// TIA Portal project "OpenLibraryExample" (V13) (continued)
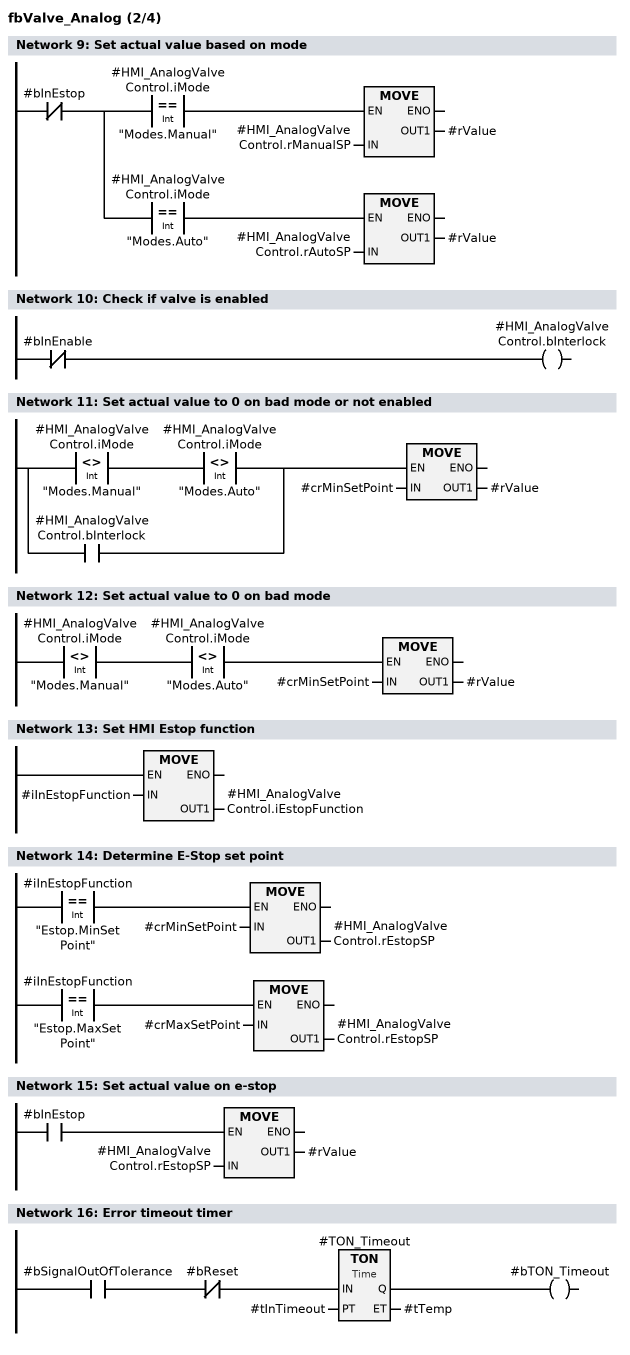
   RUNG wire#powerrail
      I_Contact( #bInEstop )
      wire#w1
      { S7_Templates := "SrcType := Int" } EQ_Contact(in1 := #HMI_AnalogValveControl.iMode, in2 := "Modes.Manual")
      { S7_GenerateENO := "TRUE" } Move(in := #HMI_AnalogValveControl.rManualSP, out1 => #rValue)
   END_RUNG
   RUNG wire#w1
      { S7_Templates := "SrcType := Int" } EQ_Contact(in1 := #HMI_AnalogValveControl.iMode, in2 := "Modes.Auto")
      { S7_GenerateENO := "TRUE" } Move(in := #HMI_AnalogValveControl.rAutoSP, out1 => #rValue)
   END_RUNG
   // the same network as SCL:
   IF NOT #bInEstop AND (#HMI_AnalogValveControl.iMode = "Modes.Manual") THEN
       #rValue := #HMI_AnalogValveControl.rManualSP;
   END_IF;
   IF NOT #bInEstop AND (#HMI_AnalogValveControl.iMode = "Modes.Auto") THEN
       #rValue := #HMI_AnalogValveControl.rAutoSP;
   END_IF;
END_REGION

REGION Network 10: Check if valve is enabled
   RUNG wire#powerrail
      I_Contact( #bInEnable )
      Coil( #HMI_AnalogValveControl.bInterlock )
   END_RUNG
   // the same network as SCL:
   #HMI_AnalogValveControl.bInterlock := NOT #bInEnable;
END_REGION

REGION Network 11: Set actual value to 0 on bad mode or not enabled
   RUNG wire#powerrail
      { S7_Templates := "SrcType := Int" } NE_Contact(in1 := #HMI_AnalogValveControl.iMode, in2 := "Modes.Manual")
      { S7_Templates := "SrcType := Int" } NE_Contact(in1 := #HMI_AnalogValveControl.iMode, in2 := "Modes.Auto")
      wire#w1
      { S7_GenerateENO := "TRUE" } Move(in := #crMinSetPoint, out1 => #rValue)
   END_RUNG
   RUNG wire#powerrail
      Contact( #HMI_AnalogValveControl.bInterlock )
   END_RUNG wire#w1
   // the same network as SCL:
   IF ((#HMI_AnalogValveControl.iMode <> "Modes.Manual") AND (#HMI_AnalogValveControl.iMode <> "Modes.Auto")) OR #HMI_AnalogValveControl.bInterlock THEN
       #rValue := #crMinSetPoint;
   END_IF;
END_REGION

REGION Network 12: Set actual value to 0 on bad mode
   RUNG wire#powerrail
      { S7_Templates := "SrcType := Int" } NE_Contact(in1 := #HMI_AnalogValveControl.iMode, in2 := "Modes.Manual")
      { S7_Templates := "SrcType := Int" } NE_Contact(in1 := #HMI_AnalogValveControl.iMode, in2 := "Modes.Auto")
      { S7_GenerateENO := "TRUE" } Move(in := #crMinSetPoint, out1 => #rValue)
   END_RUNG
   // the same network as SCL:
   IF (#HMI_AnalogValveControl.iMode <> "Modes.Manual") AND (#HMI_AnalogValveControl.iMode <> "Modes.Auto") THEN
       #rValue := #crMinSetPoint;
   END_IF;
END_REGION

REGION Network 13: Set HMI Estop function
   RUNG wire#powerrail
      Move(in := #iInEstopFunction, out1 => #HMI_AnalogValveControl.iEstopFunction)
   END_RUNG
   // the same network as SCL:
   #HMI_AnalogValveControl.iEstopFunction := #iInEstopFunction;
END_REGION

REGION Network 14: Determine E-Stop set point
   RUNG wire#powerrail
      { S7_Templates := "SrcType := Int" } EQ_Contact(in1 := #iInEstopFunction, in2 := "Estop.MinSetPoint")
      { S7_GenerateENO := "TRUE" } Move(in := #crMinSetPoint, out1 => #HMI_AnalogValveControl.rEstopSP)
   END_RUNG
   RUNG wire#powerrail
      { S7_Templates := "SrcType := Int" } EQ_Contact(in1 := #iInEstopFunction, in2 := "Estop.MaxSetPoint")
      { S7_GenerateENO := "TRUE" } Move(in := #crMaxSetPoint, out1 => #HMI_AnalogValveControl.rEstopSP)
   END_RUNG
   // the same network as SCL:
   IF #iInEstopFunction = "Estop.MinSetPoint" THEN
       #HMI_AnalogValveControl.rEstopSP := #crMinSetPoint;
   END_IF;
   IF #iInEstopFunction = "Estop.MaxSetPoint" THEN
       #HMI_AnalogValveControl.rEstopSP := #crMaxSetPoint;
   END_IF;
END_REGION

REGION Network 15: Set actual value on e-stop
   RUNG wire#powerrail
      Contact( #bInEstop )
      { S7_GenerateENO := "TRUE" } Move(in := #HMI_AnalogValveControl.rEstopSP, out1 => #rValue)
   END_RUNG
   // the same network as SCL:
   IF #bInEstop THEN #rValue := #HMI_AnalogValveControl.rEstopSP; END_IF;
END_REGION

REGION Network 16: Error timeout timer
   #TON_Timeout.TON(IN := #bSignalOutOfTolerance AND NOT #bReset, PT := #tInTimeout, ET => #tTemp);
   #bTON_Timeout := #TON_Timeout.Q;
END_REGION

REGION Network 17: Calculate tolerance limits
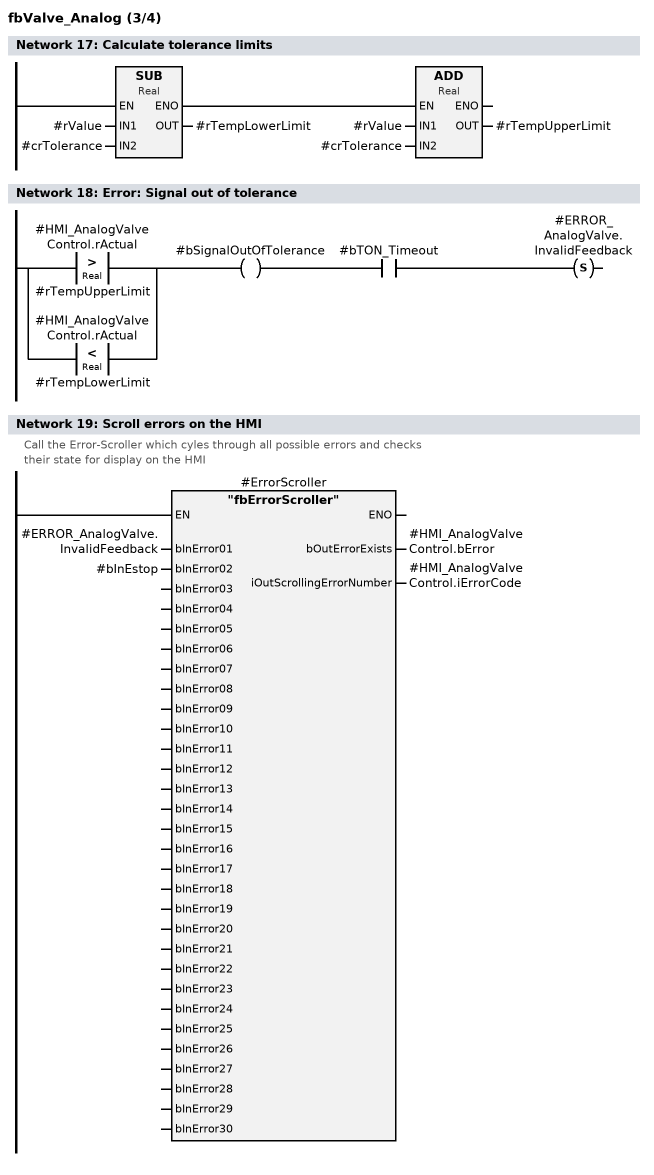
   RUNG wire#powerrail
      { S7_Templates := "SrcType := Real"; S7_GenerateENO := "TRUE" } Sub(in1 := #rValue, in2 := #crTolerance, out => #rTempLowerLimit)
      { S7_Templates := "SrcType := Real"; S7_GenerateENO := "TRUE" } Add(in1 := #rValue, in2 := #crTolerance, out => #rTempUpperLimit)
   END_RUNG
   // the same network as SCL:
   // ENO of a box is taken as its EN; it also drops when the box reports an error
   #rTempLowerLimit := #rValue - #crTolerance;
   #rTempUpperLimit := #rValue + #crTolerance;
END_REGION

REGION Network 18: Error: Signal out of tolerance
   RUNG wire#powerrail
      { S7_Templates := "SrcType := Real" } GT_Contact(in1 := #HMI_AnalogValveControl.rActual, in2 := #rTempUpperLimit)
      wire#w1
      Coil( #bSignalOutOfTolerance )
      Contact( #bTON_Timeout )
      S_Coil( #ERROR_AnalogValve.InvalidFeedback )
   END_RUNG
   RUNG wire#powerrail
      { S7_Templates := "SrcType := Real" } LT_Contact(in1 := #HMI_AnalogValveControl.rActual, in2 := #rTempLowerLimit)
   END_RUNG wire#w1
   // the same network as SCL:
   #bSignalOutOfTolerance := (#HMI_AnalogValveControl.rActual > #rTempUpperLimit) OR (#HMI_AnalogValveControl.rActual < #rTempLowerLimit);
   IF #bSignalOutOfTolerance AND #bTON_Timeout THEN #ERROR_AnalogValve.InvalidFeedback := TRUE; END_IF;
END_REGION

REGION Network 19: Scroll errors on the HMI
   // Call the Error-Scroller which cyles through all possible errors and checks 
   // their state for display on the HMI
   RUNG wire#powerrail
      #ErrorScroller(bInError01 := #ERROR_AnalogValve.InvalidFeedback, bInError02 := #bInEstop, bInError03 :=, bInError04 :=, bInError05 :=, bInError06 :=, bInError07 :=, bInError08 :=, bInError09 :=, bInError10 :=, bInError11 :=, bInError12 :=, bInError13 :=, bInError14 :=, bInError15 :=, bInError16 :=, bInError17 :=, bInError18 :=, bInError19 :=, bInError20 :=, bInError21 :=, bInError22 :=, bInError23 :=, bInError24 :=, bInError25 :=, bInError26 :=, bInError27 :=, bInError28 :=, bInError29 :=, bInError30 :=, bOutErrorExists => #HMI_AnalogValveControl.bError, iOutScrollingErrorNumber => #HMI_AnalogValveControl.iErrorCode)
   END_RUNG
   // the same network as SCL:
   #ErrorScroller(bInError01 := #ERROR_AnalogValve.InvalidFeedback,   // "fbErrorScroller"
                  bInError02 := #bInEstop,
                  bOutErrorExists => #HMI_AnalogValveControl.bError,
                  iOutScrollingErrorNumber => #HMI_AnalogValveControl.iErrorCode);
END_REGION

REGION Network 20: Set HMI status
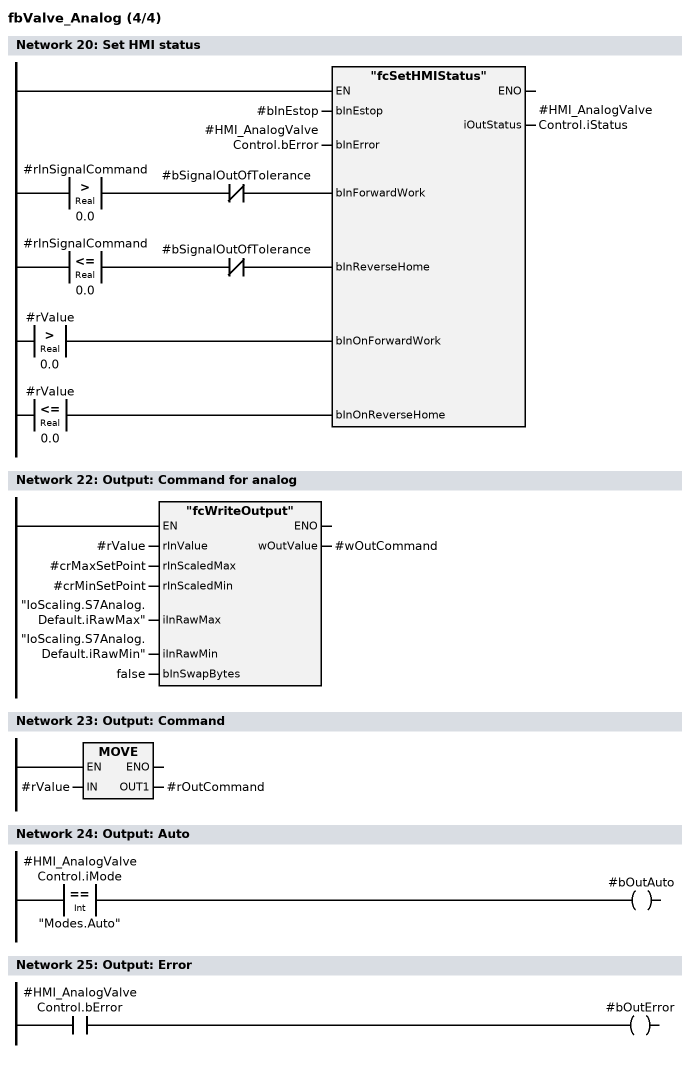
   RUNG wire#powerrail
      "fcSetHMIStatus"(bInForwardWork := wire#w1, bInReverseHome := wire#w2, bInOnForwardWork := wire#w3, bInOnReverseHome := wire#w4, bInEstop := #bInEstop, bInError := #HMI_AnalogValveControl.bError, iOutStatus => #HMI_AnalogValveControl.iStatus)
   END_RUNG
   RUNG wire#powerrail
      { S7_Templates := "SrcType := Real" } GT_Contact(in1 := #rInSignalCommand, in2 := 0.0)
      I_Contact( #bSignalOutOfTolerance )
   END_RUNG wire#w1
   RUNG wire#powerrail
      { S7_Templates := "SrcType := Real" } LE_Contact(in1 := #rInSignalCommand, in2 := 0.0)
      I_Contact( #bSignalOutOfTolerance )
   END_RUNG wire#w2
   RUNG wire#powerrail
      { S7_Templates := "SrcType := Real" } GT_Contact(in1 := #rValue, in2 := 0.0)
   END_RUNG wire#w3
   RUNG wire#powerrail
      { S7_Templates := "SrcType := Real" } LE_Contact(in1 := #rValue, in2 := 0.0)
   END_RUNG wire#w4
   // the same network as SCL:
   "fcSetHMIStatus"(bInEstop := #bInEstop,
                    bInError := #HMI_AnalogValveControl.bError,
                    bInForwardWork := (#rInSignalCommand > 0.0) AND NOT #bSignalOutOfTolerance,
                    bInReverseHome := (#rInSignalCommand <= 0.0) AND NOT #bSignalOutOfTolerance,
                    bInOnForwardWork := #rValue > 0.0,
                    bInOnReverseHome := #rValue <= 0.0,
                    iOutStatus => #HMI_AnalogValveControl.iStatus);
END_REGION

REGION Network 21: -------------------------------------------------------- Outputs --------------------------------------------------------------
END_REGION

REGION Network 22: Output: Command for analog
   RUNG wire#powerrail
      "fcWriteOutput"(rInValue := #rValue, rInScaledMax := #crMaxSetPoint, rInScaledMin := #crMinSetPoint, iInRawMax := "IoScaling.S7Analog.Default.iRawMax", iInRawMin := "IoScaling.S7Analog.Default.iRawMin", bInSwapBytes := false, wOutValue => #wOutCommand)
   END_RUNG
   // the same network as SCL:
   "fcWriteOutput"(rInValue := #rValue,
                   rInScaledMax := #crMaxSetPoint,
                   rInScaledMin := #crMinSetPoint,
                   iInRawMax := "IoScaling.S7Analog.Default.iRawMax",
                   iInRawMin := "IoScaling.S7Analog.Default.iRawMin",
                   bInSwapBytes := false,
                   wOutValue => #wOutCommand);
END_REGION

REGION Network 23: Output: Command
   RUNG wire#powerrail
      { S7_GenerateENO := "TRUE" } Move(in := #rValue, out1 => #rOutCommand)
   END_RUNG
   // the same network as SCL:
   #rOutCommand := #rValue;
END_REGION

REGION Network 24: Output: Auto
   RUNG wire#powerrail
      { S7_Templates := "SrcType := Int" } EQ_Contact(in1 := #HMI_AnalogValveControl.iMode, in2 := "Modes.Auto")
      Coil( #bOutAuto )
   END_RUNG
   // the same network as SCL:
   #bOutAuto := #HMI_AnalogValveControl.iMode = "Modes.Auto";
END_REGION

REGION Network 25: Output: Error
   RUNG wire#powerrail
      Contact( #HMI_AnalogValveControl.bError )
      Coil( #bOutError )
   END_RUNG
   // the same network as SCL:
   #bOutError := #HMI_AnalogValveControl.bError;
END_REGION
END_FUNCTION_BLOCK

FUNCTION_BLOCK "fbVFD_GSeries"   // FB120, LAD
TITLE = Controls a Siemens G120 VFD (or MicroMaster)
{ S7_Optimized_Access := 'FALSE' }
VERSION : 0.1
   VAR_TEMP   // added for the SCL form of the ladder/FBD networks
      _w1 : Bool;
      _w2 : Bool;
      _w3 : Bool;
      _w4 : Bool;
   END_VAR
BEGIN

REGION Network 1: --------------------------------------------------------- Inputs ------------------------------------------------------------------
END_REGION

REGION Network 2: Read HMI input buttons
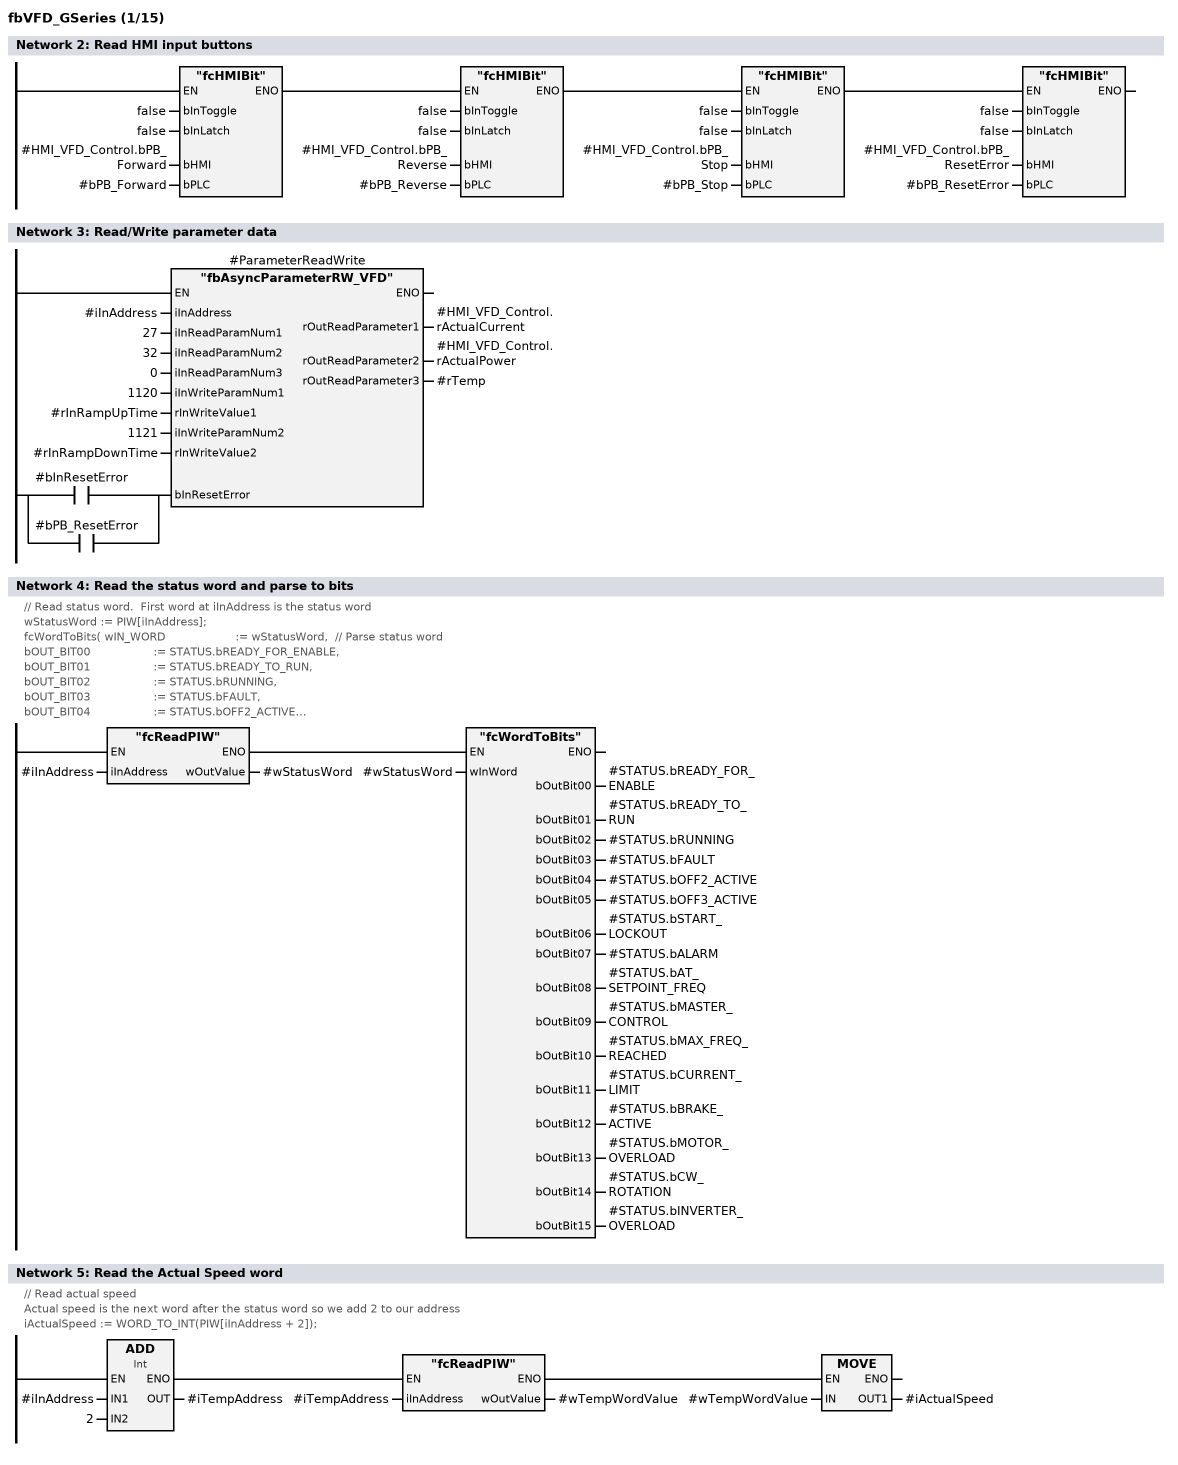
   RUNG wire#powerrail
      "fcHMIBit"(bInToggle := false, bInLatch := false, bHMI := #HMI_VFD_Control.bPB_Forward, bPLC := #bPB_Forward)
      "fcHMIBit"(bInToggle := false, bInLatch := false, bHMI := #HMI_VFD_Control.bPB_Reverse, bPLC := #bPB_Reverse)
      "fcHMIBit"(bInToggle := false, bInLatch := false, bHMI := #HMI_VFD_Control.bPB_Stop, bPLC := #bPB_Stop)
      "fcHMIBit"(bInToggle := false, bInLatch := false, bHMI := #HMI_VFD_Control.bPB_ResetError, bPLC := #bPB_ResetError)
   END_RUNG
   // the same network as SCL:
   "fcHMIBit"(bInToggle := false,
              bInLatch := false,
              bHMI := #HMI_VFD_Control.bPB_Forward,
              bPLC := #bPB_Forward,
              ENO => #_w1);
   "fcHMIBit"(EN := #_w1,
              bInToggle := false,
              bInLatch := false,
              bHMI := #HMI_VFD_Control.bPB_Reverse,
              bPLC := #bPB_Reverse,
              ENO => #_w2);
   "fcHMIBit"(EN := #_w2,
              bInToggle := false,
              bInLatch := false,
              bHMI := #HMI_VFD_Control.bPB_Stop,
              bPLC := #bPB_Stop,
              ENO => #_w3);
   IF #_w3 THEN
       "fcHMIBit"(bInToggle := false,
                  bInLatch := false,
                  bHMI := #HMI_VFD_Control.bPB_ResetError,
                  bPLC := #bPB_ResetError);
   END_IF;
END_REGION

REGION Network 3: Read/Write parameter data
   RUNG wire#powerrail
      #ParameterReadWrite(bInResetError := wire#w1, iInAddress := #iInAddress, iInReadParamNum1 := 27, iInReadParamNum2 := 32, iInReadParamNum3 := 0, iInWriteParamNum1 := 1120, rInWriteValue1 := #rInRampUpTime, iInWriteParamNum2 := 1121, rInWriteValue2 := #rInRampDownTime, rOutReadParameter1 => #HMI_VFD_Control.rActualCurrent, rOutReadParameter2 => #HMI_VFD_Control.rActualPower, rOutReadParameter3 => #rTemp)
   END_RUNG
   RUNG wire#powerrail
      Contact( #bInResetError )
   END_RUNG wire#w1
   RUNG wire#powerrail
      Contact( #bPB_ResetError )
   END_RUNG wire#w1
   // the same network as SCL:
   #ParameterReadWrite(iInAddress := #iInAddress,   // "fbAsyncParameterRW_VFD"
                       iInReadParamNum1 := 27,
                       iInReadParamNum2 := 32,
                       iInReadParamNum3 := 0,
                       iInWriteParamNum1 := 1120,
                       rInWriteValue1 := #rInRampUpTime,
                       iInWriteParamNum2 := 1121,
                       rInWriteValue2 := #rInRampDownTime,
                       bInResetError := #bInResetError OR #bPB_ResetError,
                       rOutReadParameter1 => #HMI_VFD_Control.rActualCurrent,
                       rOutReadParameter2 => #HMI_VFD_Control.rActualPower,
                       rOutReadParameter3 => #rTemp);
END_REGION

REGION Network 4: Read the status word and parse to bits
   // // Read status word.  First word at iInAddress is the status word
   // wStatusWord := PIW[iInAddress];
   // 
   // fcWordToBits( wIN_WORD                    := wStatusWord,  // Parse status word
   //                 bOUT_BIT00                  := STATUS.bREADY_FOR_ENABLE,
   //                 bOUT_BIT01                  := STATUS.bREADY_TO_RUN,
   //                 bOUT_BIT02                  := STATUS.bRUNNING,
   //                 bOUT_BIT03                  := STATUS.bFAULT,
   //                 bOUT_BIT04                  := STATUS.bOFF2_ACTIVE,
   //                 bOUT_BIT05                  := STATUS.bOFF3_ACTIVE,
   //                 bOUT_BIT06                  := STATUS.bSTART_LOCKOUT,
   //                 bOUT_BIT07                  := STATUS.bALARM,
   //                 bOUT_BIT08                  := STATUS.bAT_SETPOINT_FREQ,
   //                 bOUT_BIT09                  := STATUS.bMASTER_CONTROL,
   //                 bOUT_BIT10                  := STATUS.bMAX_FREQ_REACHED,
   //                 bOUT_BIT11                  := STATUS.bCURRENT_LIMIT,
   //                 bOUT_BIT12                  := STATUS.bBRAKE_ACTIVE,
   //                 bOUT_BIT13                  := STATUS.bMOTOR_OVERLOAD,
   //                 bOUT_BIT14                  := STATUS.bCW_ROTATION,
   //                 bOUT_BIT15                  := STATUS.bINVERTER_OVERLOAD);
   RUNG wire#powerrail
      "fcReadPIW"(iInAddress := #iInAddress, wOutValue => #wStatusWord)
      "fcWordToBits"(wInWord := #wStatusWord, bOutBit00 => #STATUS.bREADY_FOR_ENABLE, bOutBit01 => #STATUS.bREADY_TO_RUN, bOutBit02 => #STATUS.bRUNNING, bOutBit03 => #STATUS.bFAULT, bOutBit04 => #STATUS.bOFF2_ACTIVE, bOutBit05 => #STATUS.bOFF3_ACTIVE, bOutBit06 => #STATUS.bSTART_LOCKOUT, bOutBit07 => #STATUS.bALARM, bOutBit08 => #STATUS.bAT_SETPOINT_FREQ, bOutBit09 => #STATUS.bMASTER_CONTROL, bOutBit10 => #STATUS.bMAX_FREQ_REACHED, bOutBit11 => #STATUS.bCURRENT_LIMIT, bOutBit12 => #STATUS.bBRAKE_ACTIVE, bOutBit13 => #STATUS.bMOTOR_OVERLOAD, bOutBit14 => #STATUS.bCW_ROTATION, bOutBit15 => #STATUS.bINVERTER_OVERLOAD)
   END_RUNG
   // the same network as SCL:
   "fcReadPIW"(iInAddress := #iInAddress, wOutValue => #wStatusWord, ENO => #_w1);
   IF #_w1 THEN
       "fcWordToBits"(wInWord := #wStatusWord,
                      bOutBit00 => #STATUS.bREADY_FOR_ENABLE,
                      bOutBit01 => #STATUS.bREADY_TO_RUN,
                      bOutBit02 => #STATUS.bRUNNING,
                      bOutBit03 => #STATUS.bFAULT,
                      bOutBit04 => #STATUS.bOFF2_ACTIVE,
                      bOutBit05 => #STATUS.bOFF3_ACTIVE,
                      bOutBit06 => #STATUS.bSTART_LOCKOUT,
                      bOutBit07 => #STATUS.bALARM,
                      bOutBit08 => #STATUS.bAT_SETPOINT_FREQ,
                      bOutBit09 => #STATUS.bMASTER_CONTROL,
                      bOutBit10 => #STATUS.bMAX_FREQ_REACHED,
                      bOutBit11 => #STATUS.bCURRENT_LIMIT,
                      bOutBit12 => #STATUS.bBRAKE_ACTIVE,
                      bOutBit13 => #STATUS.bMOTOR_OVERLOAD,
                      bOutBit14 => #STATUS.bCW_ROTATION,
                      bOutBit15 => #STATUS.bINVERTER_OVERLOAD);
   END_IF;
END_REGION

REGION Network 5: Read the Actual Speed word
   // // Read actual speed
   // Actual speed is the next word after the status word so we add 2 to our address
   // iActualSpeed := WORD_TO_INT(PIW[iInAddress + 2]);
   RUNG wire#powerrail
      { S7_Templates := "SrcType := Int"; S7_GenerateENO := "TRUE" } Add(in1 := #iInAddress, in2 := 2, out => #iTempAddress)
      "fcReadPIW"(iInAddress := #iTempAddress, wOutValue => #wTempWordValue)
      { S7_GenerateENO := "TRUE" } Move(in := #wTempWordValue, out1 => #iActualSpeed)
   END_RUNG
   // the same network as SCL:
   // ENO of a box is taken as its EN; it also drops when the box reports an error
   #iTempAddress := #iInAddress + 2;
   "fcReadPIW"(iInAddress := #iTempAddress, wOutValue => #wTempWordValue, ENO => #_w1);
   IF #_w1 THEN #iActualSpeed := #wTempWordValue; END_IF;
END_REGION

REGION Network 6: Update the signal forward bit
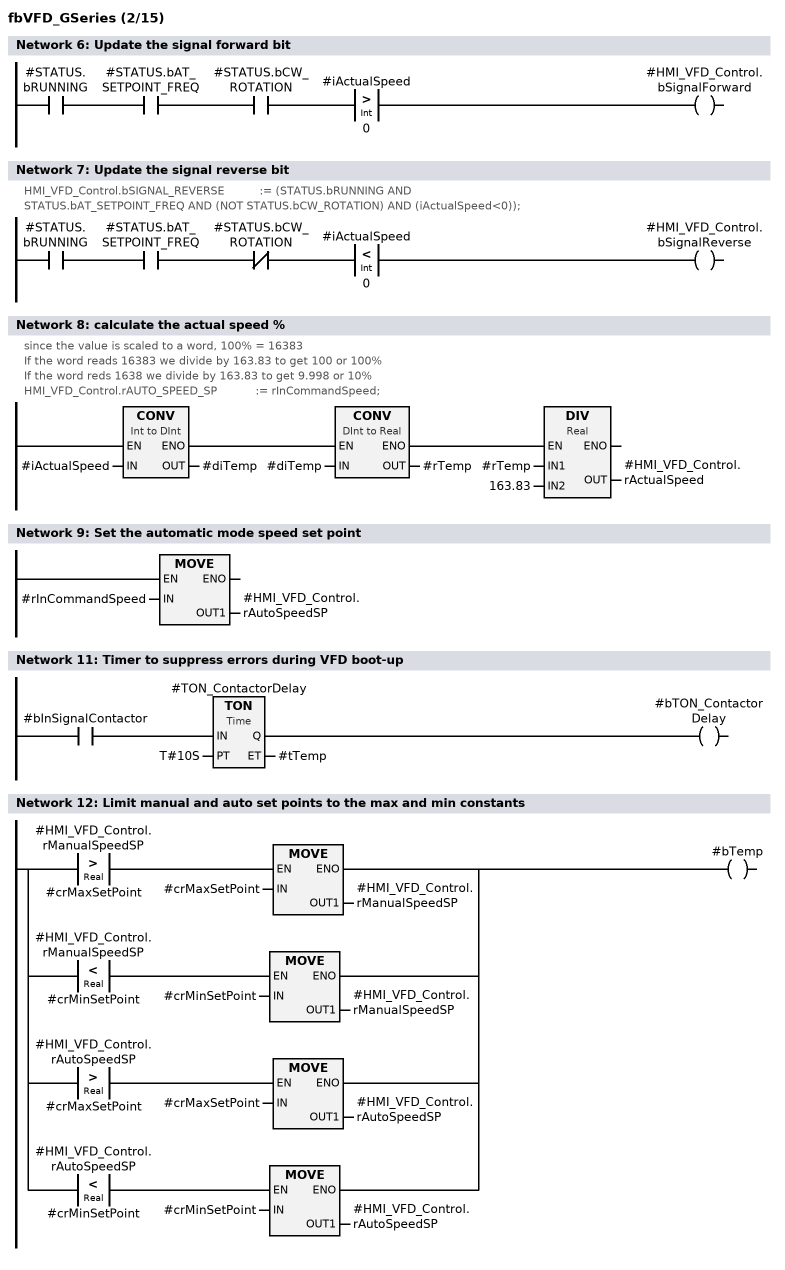
   RUNG wire#powerrail
      Contact( #STATUS.bRUNNING )
      Contact( #STATUS.bAT_SETPOINT_FREQ )
      Contact( #STATUS.bCW_ROTATION )
      { S7_Templates := "SrcType := Int" } GT_Contact(in1 := #iActualSpeed, in2 := 0)
      Coil( #HMI_VFD_Control.bSignalForward )
   END_RUNG
   // the same network as SCL:
   #HMI_VFD_Control.bSignalForward := #STATUS.bRUNNING AND #STATUS.bAT_SETPOINT_FREQ AND #STATUS.bCW_ROTATION AND (#iActualSpeed > 0);
END_REGION

REGION Network 7: Update the signal reverse bit
   // HMI_VFD_Control.bSIGNAL_REVERSE          := (STATUS.bRUNNING AND 
   // STATUS.bAT_SETPOINT_FREQ AND (NOT STATUS.bCW_ROTATION) AND (iActualSpeed<0));
   RUNG wire#powerrail
      Contact( #STATUS.bRUNNING )
      Contact( #STATUS.bAT_SETPOINT_FREQ )
      I_Contact( #STATUS.bCW_ROTATION )
      { S7_Templates := "SrcType := Int" } LT_Contact(in1 := #iActualSpeed, in2 := 0)
      Coil( #HMI_VFD_Control.bSignalReverse )
   END_RUNG
   // the same network as SCL:
   #HMI_VFD_Control.bSignalReverse := #STATUS.bRUNNING AND #STATUS.bAT_SETPOINT_FREQ AND NOT #STATUS.bCW_ROTATION AND (#iActualSpeed < 0);
END_REGION

REGION Network 8: calculate the actual speed %
   // since the value is scaled to a word, 100% = 16383
   // 
   // If the word reads 16383 we divide by 163.83 to get 100 or 100%
   // If the word reds 1638 we divide by 163.83 to get 9.998 or 10%
   // 
   // HMI_VFD_Control.rAUTO_SPEED_SP           := rInCommandSpeed;
   RUNG wire#powerrail
      { S7_Templates := "[SrcType := Int, DestType := DInt]"; S7_GenerateENO := "TRUE" } Convert(in := #iActualSpeed, out => #diTemp)
      { S7_Templates := "[SrcType := DInt, DestType := Real]"; S7_GenerateENO := "TRUE" } Convert(in := #diTemp, out => #rTemp)
      { S7_Templates := "SrcType := Real"; S7_GenerateENO := "TRUE" } Div(in1 := #rTemp, in2 := 163.83, out => #HMI_VFD_Control.rActualSpeed)
   END_RUNG
   // the same network as SCL:
   // ENO of a box is taken as its EN; it also drops when the box reports an error
   #diTemp := INT_TO_DINT(#iActualSpeed);
   #rTemp := DINT_TO_REAL(#diTemp);
   #HMI_VFD_Control.rActualSpeed := #rTemp / 163.83;
END_REGION

REGION Network 9: Set the automatic mode speed set point
   RUNG wire#powerrail
      { S7_GenerateENO := "TRUE" } Move(in := #rInCommandSpeed, out1 => #HMI_VFD_Control.rAutoSpeedSP)
   END_RUNG
   // the same network as SCL:
   #HMI_VFD_Control.rAutoSpeedSP := #rInCommandSpeed;
END_REGION

REGION Network 10: --------------------------------------------------- Control Logic ------------------------------------------------------------
END_REGION

REGION Network 11: Timer to suppress errors during VFD boot-up
   #TON_ContactorDelay.TON(IN := #bInSignalContactor, PT := T#10S, ET => #tTemp);
   #bTON_ContactorDelay := #TON_ContactorDelay.Q;
END_REGION

REGION Network 12: Limit manual and auto set points to the max and min constants
   RUNG wire#powerrail
      { S7_Templates := "SrcType := Real" } GT_Contact(in1 := #HMI_VFD_Control.rManualSpeedSP, in2 := #crMaxSetPoint)
      { S7_GenerateENO := "TRUE" } Move(in := #crMaxSetPoint, out1 => #HMI_VFD_Control.rManualSpeedSP)
      wire#w1
      Coil( #bTemp )
   END_RUNG
   RUNG wire#powerrail
      { S7_Templates := "SrcType := Real" } LT_Contact(in1 := #HMI_VFD_Control.rManualSpeedSP, in2 := #crMinSetPoint)
      { S7_GenerateENO := "TRUE" } Move(in := #crMinSetPoint, out1 => #HMI_VFD_Control.rManualSpeedSP)
   END_RUNG wire#w1
   RUNG wire#powerrail
      { S7_Templates := "SrcType := Real" } GT_Contact(in1 := #HMI_VFD_Control.rAutoSpeedSP, in2 := #crMaxSetPoint)
      { S7_GenerateENO := "TRUE" } Move(in := #crMaxSetPoint, out1 => #HMI_VFD_Control.rAutoSpeedSP)
   END_RUNG wire#w1
   RUNG wire#powerrail
      { S7_Templates := "SrcType := Real" } LT_Contact(in1 := #HMI_VFD_Control.rAutoSpeedSP, in2 := #crMinSetPoint)
      { S7_GenerateENO := "TRUE" } Move(in := #crMinSetPoint, out1 => #HMI_VFD_Control.rAutoSpeedSP)
   END_RUNG wire#w1
   // the same network as SCL:
   // ENO of a box is taken as its EN; it also drops when the box reports an error
   #_w1 := #HMI_VFD_Control.rManualSpeedSP > #crMaxSetPoint;
   IF #_w1 THEN #HMI_VFD_Control.rManualSpeedSP := #crMaxSetPoint; END_IF;
   #_w2 := #HMI_VFD_Control.rManualSpeedSP < #crMinSetPoint;
   IF #_w2 THEN #HMI_VFD_Control.rManualSpeedSP := #crMinSetPoint; END_IF;
   #_w3 := #HMI_VFD_Control.rAutoSpeedSP > #crMaxSetPoint;
   IF #_w3 THEN #HMI_VFD_Control.rAutoSpeedSP := #crMaxSetPoint; END_IF;
   #_w4 := #HMI_VFD_Control.rAutoSpeedSP < #crMinSetPoint;
   IF #_w4 THEN #HMI_VFD_Control.rAutoSpeedSP := #crMinSetPoint; END_IF;
   #bTemp := #_w1 OR #_w2 OR #_w3 OR #_w4;
END_REGION

REGION Network 13: Reset errors
   // Clear all errors
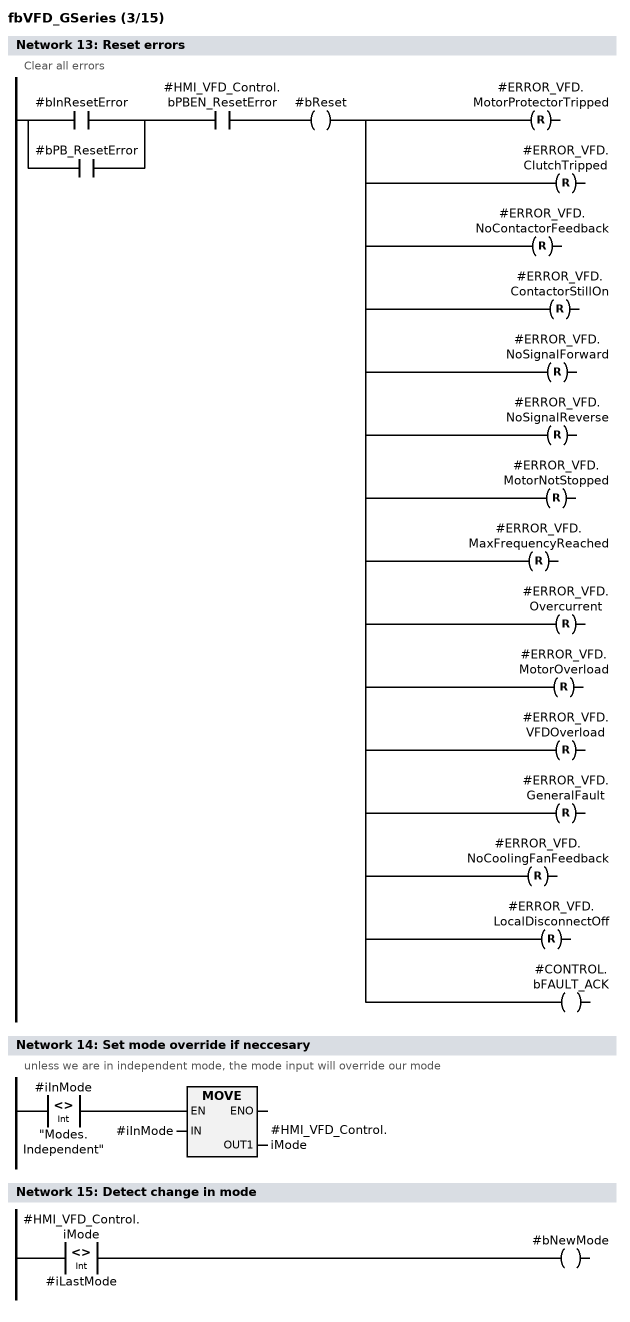
   RUNG wire#powerrail
      Contact( #bInResetError )
      wire#w1
      Contact( #HMI_VFD_Control.bPBEN_ResetError )
      Coil( #bReset )
      wire#w2
      R_Coil( #ERROR_VFD.MotorProtectorTripped )
   END_RUNG
   RUNG wire#powerrail
      Contact( #bPB_ResetError )
   END_RUNG wire#w1
   RUNG wire#w2
      R_Coil( #ERROR_VFD.ClutchTripped )
   END_RUNG
   RUNG wire#w2
      R_Coil( #ERROR_VFD.NoContactorFeedback )
   END_RUNG
   RUNG wire#w2
      R_Coil( #ERROR_VFD.ContactorStillOn )
   END_RUNG
   RUNG wire#w2
      R_Coil( #ERROR_VFD.NoSignalForward )
   END_RUNG
   RUNG wire#w2
      R_Coil( #ERROR_VFD.NoSignalReverse )
   END_RUNG
   RUNG wire#w2
      R_Coil( #ERROR_VFD.MotorNotStopped )
   END_RUNG
   RUNG wire#w2
      R_Coil( #ERROR_VFD.MaxFrequencyReached )
   END_RUNG
   RUNG wire#w2
      R_Coil( #ERROR_VFD.Overcurrent )
   END_RUNG
   RUNG wire#w2
      R_Coil( #ERROR_VFD.MotorOverload )
   END_RUNG
   RUNG wire#w2
      R_Coil( #ERROR_VFD.VFDOverload )
   END_RUNG
   RUNG wire#w2
      R_Coil( #ERROR_VFD.GeneralFault )
   END_RUNG
   RUNG wire#w2
      R_Coil( #ERROR_VFD.NoCoolingFanFeedback )
   END_RUNG
   RUNG wire#w2
      R_Coil( #ERROR_VFD.LocalDisconnectOff )
   END_RUNG
   RUNG wire#w2
      Coil( #CONTROL.bFAULT_ACK )
   END_RUNG
   // the same network as SCL:
   #bReset := (#bInResetError OR #bPB_ResetError) AND #HMI_VFD_Control.bPBEN_ResetError;
   IF #bReset THEN
       #ERROR_VFD.MotorProtectorTripped := FALSE;
       #ERROR_VFD.ClutchTripped := FALSE;
       #ERROR_VFD.NoContactorFeedback := FALSE;
       #ERROR_VFD.ContactorStillOn := FALSE;
       #ERROR_VFD.NoSignalForward := FALSE;
       #ERROR_VFD.NoSignalReverse := FALSE;
       #ERROR_VFD.MotorNotStopped := FALSE;
       #ERROR_VFD.MaxFrequencyReached := FALSE;
       #ERROR_VFD.Overcurrent := FALSE;
       #ERROR_VFD.MotorOverload := FALSE;
       #ERROR_VFD.VFDOverload := FALSE;
       #ERROR_VFD.GeneralFault := FALSE;
       #ERROR_VFD.NoCoolingFanFeedback := FALSE;
       #ERROR_VFD.LocalDisconnectOff := FALSE;
   END_IF;
   #CONTROL.bFAULT_ACK := #bReset;
END_REGION

REGION Network 14: Set mode override if neccesary
   // unless we are in independent mode, the mode input will override our mode
   RUNG wire#powerrail
      { S7_Templates := "SrcType := Int" } NE_Contact(in1 := #iInMode, in2 := "Modes.Independent")
      { S7_GenerateENO := "TRUE" } Move(in := #iInMode, out1 => #HMI_VFD_Control.iMode)
   END_RUNG
   // the same network as SCL:
   IF #iInMode <> "Modes.Independent" THEN #HMI_VFD_Control.iMode := #iInMode; END_IF;
END_REGION

REGION Network 15: Detect change in mode
   RUNG wire#powerrail
      { S7_Templates := "SrcType := Int" } NE_Contact(in1 := #HMI_VFD_Control.iMode, in2 := #iLastMode)
      Coil( #bNewMode )
   END_RUNG
   // the same network as SCL:
   #bNewMode := #HMI_VFD_Control.iMode <> #iLastMode;
END_REGION

REGION Network 16: Keep track of last mode
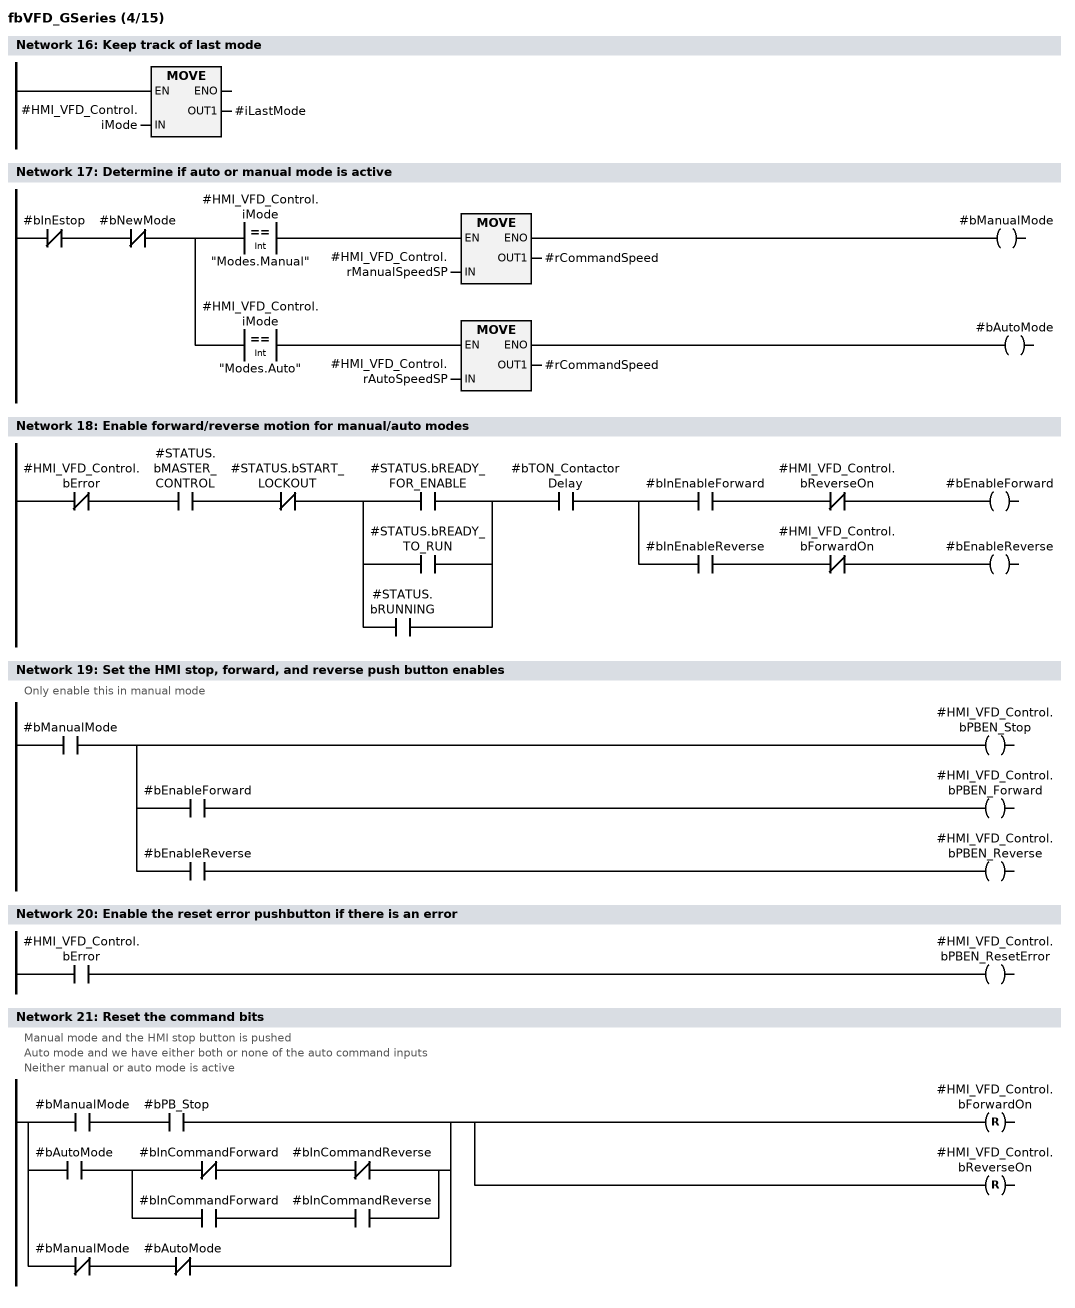
   RUNG wire#powerrail
      { S7_GenerateENO := "TRUE" } Move(in := #HMI_VFD_Control.iMode, out1 => #iLastMode)
   END_RUNG
   // the same network as SCL:
   #iLastMode := #HMI_VFD_Control.iMode;
END_REGION

REGION Network 17: Determine if auto or manual mode is active
   RUNG wire#powerrail
      I_Contact( #bInEstop )
      I_Contact( #bNewMode )
      wire#w1
      { S7_Templates := "SrcType := Int" } EQ_Contact(in1 := #HMI_VFD_Control.iMode, in2 := "Modes.Manual")
      { S7_GenerateENO := "TRUE" } Move(in := #HMI_VFD_Control.rManualSpeedSP, out1 => #rCommandSpeed)
      Coil( #bManualMode )
   END_RUNG
   RUNG wire#w1
      { S7_Templates := "SrcType := Int" } EQ_Contact(in1 := #HMI_VFD_Control.iMode, in2 := "Modes.Auto")
      { S7_GenerateENO := "TRUE" } Move(in := #HMI_VFD_Control.rAutoSpeedSP, out1 => #rCommandSpeed)
      Coil( #bAutoMode )
   END_RUNG
   // the same network as SCL:
   // ENO of a box is taken as its EN; it also drops when the box reports an error
   #_w1 := NOT #bInEstop AND NOT #bNewMode;
   #_w2 := #_w1 AND (#HMI_VFD_Control.iMode = "Modes.Manual");
   IF #_w2 THEN #rCommandSpeed := #HMI_VFD_Control.rManualSpeedSP; END_IF;
   #bManualMode := #_w2;
   #_w3 := #_w1 AND (#HMI_VFD_Control.iMode = "Modes.Auto");
   IF #_w3 THEN #rCommandSpeed := #HMI_VFD_Control.rAutoSpeedSP; END_IF;
   #bAutoMode := #_w3;
END_REGION

REGION Network 18: Enable forward/reverse motion for manual/auto modes
   RUNG wire#powerrail
      I_Contact( #HMI_VFD_Control.bError )
      Contact( #STATUS.bMASTER_CONTROL )
      I_Contact( #STATUS.bSTART_LOCKOUT )
      wire#w1
      Contact( #STATUS.bREADY_FOR_ENABLE )
      wire#w2
      Contact( #bTON_ContactorDelay )
      wire#w3
      Contact( #bInEnableForward )
      I_Contact( #HMI_VFD_Control.bReverseOn )
      Coil( #bEnableForward )
   END_RUNG
   RUNG wire#w1
      Contact( #STATUS.bREADY_TO_RUN )
   END_RUNG wire#w2
   RUNG wire#w1
      Contact( #STATUS.bRUNNING )
   END_RUNG wire#w2
   RUNG wire#w3
      Contact( #bInEnableReverse )
      I_Contact( #HMI_VFD_Control.bForwardOn )
      Coil( #bEnableReverse )
   END_RUNG
   // the same network as SCL:
   #_w1 := NOT #HMI_VFD_Control.bError AND #STATUS.bMASTER_CONTROL AND NOT #STATUS.bSTART_LOCKOUT AND (#STATUS.bREADY_FOR_ENABLE OR #STATUS.bREADY_TO_RUN OR #STATUS.bRUNNING) AND #bTON_ContactorDelay;
   #bEnableForward := #_w1 AND #bInEnableForward AND NOT #HMI_VFD_Control.bReverseOn;
   #bEnableReverse := #_w1 AND #bInEnableReverse AND NOT #HMI_VFD_Control.bForwardOn;
END_REGION

REGION Network 19: Set the HMI stop, forward, and reverse push button enables
   // Only enable this in manual mode
   RUNG wire#powerrail
      Contact( #bManualMode )
      wire#w1
      Coil( #HMI_VFD_Control.bPBEN_Stop )
   END_RUNG
   RUNG wire#w1
      Contact( #bEnableForward )
      Coil( #HMI_VFD_Control.bPBEN_Forward )
   END_RUNG
   RUNG wire#w1
      Contact( #bEnableReverse )
      Coil( #HMI_VFD_Control.bPBEN_Reverse )
   END_RUNG
   // the same network as SCL:
   #HMI_VFD_Control.bPBEN_Stop := #bManualMode;
   #HMI_VFD_Control.bPBEN_Forward := #bManualMode AND #bEnableForward;
   #HMI_VFD_Control.bPBEN_Reverse := #bManualMode AND #bEnableReverse;
END_REGION

REGION Network 20: Enable the reset error pushbutton if there is an error
   RUNG wire#powerrail
      Contact( #HMI_VFD_Control.bError )
      Coil( #HMI_VFD_Control.bPBEN_ResetError )
   END_RUNG
   // the same network as SCL:
   #HMI_VFD_Control.bPBEN_ResetError := #HMI_VFD_Control.bError;
END_REGION

REGION Network 21: Reset the command bits
   // Manual mode and the HMI stop button is pushed
   // Auto mode and we have either both or none of the auto command inputs
   // Neither manual or auto mode is active
   RUNG wire#powerrail
      Contact( #bManualMode )
      Contact( #bPB_Stop )
      wire#w1
      R_Coil( #HMI_VFD_Control.bForwardOn )
   END_RUNG
   RUNG wire#powerrail
      Contact( #bAutoMode )
      wire#w2
      I_Contact( #bInCommandForward )
      I_Contact( #bInCommandReverse )
   END_RUNG wire#w1
   RUNG wire#w2
      Contact( #bInCommandForward )
      Contact( #bInCommandReverse )
   END_RUNG wire#w1
   RUNG wire#powerrail
      I_Contact( #bManualMode )
      I_Contact( #bAutoMode )
   END_RUNG wire#w1
   RUNG wire#w1
      R_Coil( #HMI_VFD_Control.bReverseOn )
   END_RUNG
   // the same network as SCL:
   IF (#bManualMode AND #bPB_Stop) OR (#bAutoMode AND ((NOT #bInCommandForward AND NOT #bInCommandReverse) OR (#bInCommandForward AND #bInCommandReverse))) OR (NOT #bManualMode AND NOT #bAutoMode) THEN
       #HMI_VFD_Control.bForwardOn := FALSE;
       #HMI_VFD_Control.bReverseOn := FALSE;
   END_IF;
END_REGION

REGION Network 22: Start forward request
   // Manual mode and only a start forward button is pressed and enabled
   // Auto mode when we receive a auto command and it is enabled